                 // Check if line contains FOR token
                 IF FIND(IN1 := #lineBuffer.lines[#lineBuffer.pointers.retrievePointer].content, IN2 := #statKeyToken.tokenFor) <> 0 THEN
                   // Tokenize line where retrieve pointer is pointing at
                   #tempReturnVal := "LKinLang_TokenizeSlot"(lastIndexOfMerger := #statLastIndexOfMerger,
                                                             lineNumber := #lineBuffer.lines[#lineBuffer.pointers.retrievePointer].number,
                                                             line := #lineBuffer.lines[#lineBuffer.pointers.retrievePointer].content,
                                                             separators := #statSeparators,
                                                             mergers := #statMergers,
                                                             preprocessorConfig := #preProcessConfig,
                                                             tokenizedLine => #statTokenizedLine,
                                                             errorString := #statErrorString);

                   // Check if line has content
                   IF #statTokenizedLine.numberOfToken > 0 THEN
                     // Check if line starts with FOR token
                     IF #statTokenizedLine.lineToken[#statTokenizedLine.numberOfToken] = #statKeyToken.tokenFor THEN
                       // Increase array index
                       #statHierarchicLevel.numberOfLevels += 1;
                       // Check if index is ok
                       IF #statHierarchicLevel.numberOfLevels <= "LKINLANG_NUMBER_OF_HIERARCHICLEVEL" THEN
                         // Increase hierarchic level
                         #statHierarchicLevel.currentLevel += 1;
                         // Store entry
                         #statHierarchicLevel.levels[#statHierarchicLevel.numberOfLevels].level := #statHierarchicLevel.currentLevel;
                         #statHierarchicLevel.levels[#statHierarchicLevel.numberOfLevels].lineNumber := #statTokenizedLine.lineNo;
                         #statHierarchicLevel.levels[#statHierarchicLevel.numberOfLevels].type := "LKINLANG_ENTRY_TYPE_FOR"; // Type for FOR
                       ELSE
                         // Error hierarchic level array overflow
                         #statStatus := #ERR_HIERARCHIC_LEVEL_LIST;
                         #statStateIntern := #STATE_ERROR;
                         #statErrorString := CONCAT(IN1 := #statErrorString, IN2 := 'Error: Maximum array index of hierarchic level reached');
                         #statErrorString := CONCAT(IN1 := #statErrorString, IN2 := ' in line: ');
                         #statErrorString := CONCAT(IN1 := #statErrorString, IN2 := UDINT_TO_STRING(#statTokenizedLine.lineNo));
                       END_IF;
                     END_IF;
                   END_IF;
                 END_IF;

                 // Check if line contains ENDFOR token
                 IF FIND(IN1 := #lineBuffer.lines[#lineBuffer.pointers.retrievePointer].content, IN2 := #statKeyToken.tokenEndFor) <> 0 THEN
                   // Tokenize line where retrieve pointer is pointing at
                   #tempReturnVal := "LKinLang_TokenizeSlot"(lastIndexOfMerger := #statLastIndexOfMerger,
                                                             lineNumber := #lineBuffer.lines[#lineBuffer.pointers.retrievePointer].number,
                                                             line := #lineBuffer.lines[#lineBuffer.pointers.retrievePointer].content,
                                                             separators := #statSeparators,
                                                             mergers := #statMergers,
                                                             preprocessorConfig := #preProcessConfig,
                                                             tokenizedLine => #statTokenizedLine,
                                                             errorString := #statErrorString);

                   // Check if line has content
                   IF #statTokenizedLine.numberOfToken > 0 THEN
                     // Check if line starts with ENDFOR token
                     IF #statTokenizedLine.lineToken[#statTokenizedLine.numberOfToken] = #statKeyToken.tokenEndFor THEN
                       // Increase array index
                       #statHierarchicLevel.numberOfLevels += 1;
                       // Check if index is ok
                       IF #statHierarchicLevel.numberOfLevels <= "LKINLANG_NUMBER_OF_HIERARCHICLEVEL" THEN
                         // Store entry
                         #statHierarchicLevel.levels[#statHierarchicLevel.numberOfLevels].level := #statHierarchicLevel.currentLevel;
                         #statHierarchicLevel.levels[#statHierarchicLevel.numberOfLevels].lineNumber := #statTokenizedLine.lineNo;
                         #statHierarchicLevel.levels[#statHierarchicLevel.numberOfLevels].type := "LKINLANG_ENTRY_TYPE_ENDFOR"; // Type for ENDFOR

                         // Decrease hierarchic level
                         #statHierarchicLevel.currentLevel -= 1;
                       ELSE
                         // Error hierarchic level array overflow
                         #statStatus := #ERR_HIERARCHIC_LEVEL_LIST;
                         #statStateIntern := #STATE_ERROR;
                         #statErrorString := CONCAT(IN1 := #statErrorString, IN2 := 'Error: Maximum array index of hierarchic level reached');
                         #statErrorString := CONCAT(IN1 := #statErrorString, IN2 := ' in line: ');
                         #statErrorString := CONCAT(IN1 := #statErrorString, IN2 := UDINT_TO_STRING(#statTokenizedLine.lineNo));
                       END_IF;
                     END_IF;
                   END_IF;
                 END_IF;
               END_REGION GET_HIERARCHIC_LEVEL

               // Check if error occurred and exit reapeat
               IF #statStateIntern = #STATE_ERROR THEN
                 EXIT;
               END_IF;

               // ------------------------------------------------------------------------------------------
               // Search labels in program
               // ------------------------------------------------------------------------------------------
               // Check if LABEL key token is in line 
               // YES: Tokenize line
               // NO: next line
               REGION GENERATE_LABEL_LIST
                 // Check if line contains LABEL token
                 IF FIND(IN1 := #lineBuffer.lines[#lineBuffer.pointers.retrievePointer].content, IN2 := #statKeyToken.tokenJumpTarget) <> 0 THEN

                   // Tokenize line where retrieve pointer is pointing at
                   #tempReturnVal := "LKinLang_TokenizeSlot"(lastIndexOfMerger := #statLastIndexOfMerger,
                                                             lineNumber := #lineBuffer.lines[#lineBuffer.pointers.retrievePointer].number,
                                                             line := #lineBuffer.lines[#lineBuffer.pointers.retrievePointer].content,
                                                             separators := #statSeparators,
                                                             mergers := #statMergers,
                                                             preprocessorConfig := #preProcessConfig,
                                                             tokenizedLine => #statTokenizedLine,
                                                             errorString := #statErrorString);

                   // Check for error while tokenizing
                   IF #tempReturnVal <> 0 THEN
                     // Error while tokenizing
                     #statStatus := #ERR_TOKENIZING;
                     #statStateIntern := #STATE_ERROR;
                     EXIT;
                   END_IF;


                   // Check if line has content
                   IF #statTokenizedLine.numberOfToken > 0 THEN // Line has content --> Parse
                     // Go to ParseLine state if tokenizing was successful
                     // Check if line starts with 'LABEL'
                     IF #statTokenizedLine.lineToken[#statTokenizedLine.numberOfToken] = #statKeyToken.tokenJumpTarget THEN
                       // Check if line contains exactly 3 tokens
                       // Definition:
                       // [1] "myLabel"
                       // [2] " "
                       // [3] "LABEL"
                       IF #statTokenizedLine.numberOfToken = 3 THEN
                         IF #statTokenizedLine.lineToken[#statTokenizedLine.numberOfToken - 1] = ' ' // second token must be space
                           AND NOT "LKinLang_IsTokenNumberInclSign"(#statTokenizedLine.lineToken[#statTokenizedLine.numberOfToken - 2]) // first token must not be a number
                         THEN
                           // correct label definition 
                           // Check labelList if label already exists
                           FOR #tempCounter := 1 TO #statLabelList.numberOfLabels DO
                             IF #statLabelList.labels[#tempCounter].labelName = #statTokenizedLine.lineToken[#statTokenizedLine.numberOfToken - 2] THEN
                               // Label already exists in other line
                               // Throw error
                               #statStatus := #ERR_LABEL_LIST;
                               #statStateIntern := #STATE_ERROR;
                               #statErrorString := CONCAT(IN1 := #statErrorString, IN2 := ';Error: Label is not unique');
                               #statErrorString := CONCAT(IN1 := #statErrorString, IN2 := ' in line: ');
                               #statErrorString := CONCAT(IN1 := #statErrorString, IN2 := UDINT_TO_STRING(#statTokenizedLine.lineNo));
                               EXIT;
                             END_IF;
                           END_FOR;

                           // Check if error was set in for loop
                           // --> Abort repeat loop 
                           IF #statStateIntern = #STATE_ERROR THEN
                             EXIT;
                           END_IF;

                           // Check if name is a keyword
                           IF "LKinLang_IsTokenKeyWord"(token := #statTokenizedLine.lineToken[#statTokenizedLine.numberOfToken - 2], keyToken := #statKeyToken) THEN
                             // Error: Label name can not be a keyword
                             #statStatus := #ERR_LABEL_LIST;
                             #statStateIntern := #STATE_ERROR;
                             #statErrorString := CONCAT(IN1 := #statErrorString, IN2 := 'Error: Label name must not be a keyword');
                             #statErrorString := CONCAT(IN1 := #statErrorString, IN2 := '; Line: ');
                             #statErrorString := CONCAT(IN1 := #statErrorString, IN2 := UDINT_TO_STRING(#statTokenizedLine.lineNo));
                             EXIT;
                           END_IF;

                           // Check if name is a parameter 
                           FOR #tempVarIndex := 1 TO "LKINLANG_MAX_NUMBER_OF_PARAMETERS" DO
                             IF #statParameterLookUpTable[#tempVarIndex].parameterNameString = #statTokenizedLine.lineToken[#statTokenizedLine.numberOfToken - 2] THEN
                               // Error: Label name can not be a parameter
                               #statStatus := #ERR_LABEL_LIST;
                               #statStateIntern := #STATE_ERROR;
                               #statErrorString := CONCAT(IN1 := #statErrorString, IN2 := 'Error: Label name must not be a keyword');
                               #statErrorString := CONCAT(IN1 := #statErrorString, IN2 := '; Line: ');
                               #statErrorString := CONCAT(IN1 := #statErrorString, IN2 := UDINT_TO_STRING(#statTokenizedLine.lineNo));
                               EXIT;
                             END_IF;
                           END_FOR;

                           // Check if error was set in for loop
                           // --> Abort repeat loop 
                           IF #statStateIntern = #STATE_ERROR THEN
                             EXIT;
                           END_IF;

                           // Check if the number of labels is ok 
                           IF #statLabelList.numberOfLabels >= "LKINLANG_NUMBER_OF_LABELS" THEN
                             // No more space in labelList
                             // Throw error 
                             #statStatus := #ERR_LABEL_LIST;
                             #statStateIntern := #STATE_ERROR;
                             #statErrorString := CONCAT(IN1 := #statErrorString, IN2 := ';Error: Maximum number of labels reached');
                             #statErrorString := CONCAT(IN1 := #statErrorString, IN2 := ' in line: ');
                             #statErrorString := CONCAT(IN1 := #statErrorString, IN2 := UDINT_TO_STRING(#statTokenizedLine.lineNo));
                             EXIT;
                           END_IF;

                           IF #statStateIntern <> #STATE_ERROR THEN
                             // Increment number of labels
                             #statLabelList.numberOfLabels += 1;
                             // Set the label info
                             #statLabelList.labels[#statLabelList.numberOfLabels].labelName := #statTokenizedLine.lineToken[#statTokenizedLine.numberOfToken - 2];
                             #statLabelList.labels[#statLabelList.numberOfLabels].lineNumber := #statTokenizedLine.lineNo;
                             IF #statHierarchicLevel.numberOfLevels > 0 THEN
                               #statLabelList.labels[#statLabelList.numberOfLabels].hierarchicLevel := #statHierarchicLevel.levels[#statHierarchicLevel.numberOfLevels].level;
                             ELSE
                               #statLabelList.labels[#statLabelList.numberOfLabels].hierarchicLevel := 0;
                             END_IF;
                           ELSE
                             // Error was set already set
                             // Do nothing
                             ;
                           END_IF;

                         ELSE
                           // Wrong label definition --> No space or correct name
                           // Throw error
                           #statStatus := #ERR_LABEL_LIST;
                           #statStateIntern := #STATE_ERROR;
                           #statErrorString := CONCAT(IN1 := #statErrorString, IN2 := ';Error: Invalid label definition');
                           #statErrorString := CONCAT(IN1 := #statErrorString, IN2 := ' in line: ');
                           #statErrorString := CONCAT(IN1 := #statErrorString, IN2 := UDINT_TO_STRING(#statTokenizedLine.lineNo));
                           EXIT;
                         END_IF;
                       ELSE
                         // Wrong label definition --> Not 3 token
                         // Throw error
                         #statStatus := #ERR_LABEL_LIST;
                         #statStateIntern := #STATE_ERROR;
                         #statErrorString := CONCAT(IN1 := #statErrorString, IN2 := ';Error: Invalid label definition');
                         #statErrorString := CONCAT(IN1 := #statErrorString, IN2 := ' in line: ');
                         #statErrorString := CONCAT(IN1 := #statErrorString, IN2 := UDINT_TO_STRING(#statTokenizedLine.lineNo));
                         EXIT;
                       END_IF;

                     ELSE
                       ;// Not a label definition
                     END_IF;
                   ELSE
                     ; // Line is empty --> Tokenize next Line
                   END_IF;
                 END_IF;
               END_REGION GENERATE_LABEL_LIST

               // ------------------------------------------------------------------------------------------
               // Search sub programs
               // ------------------------------------------------------------------------------------------
               // Check if SUB key token is in line 
               REGION SUB_PROGRAM
                 // Check if line contains SUB token
                 IF FIND(IN1 := #lineBuffer.lines[#lineBuffer.pointers.retrievePointer].content, IN2 := #statKeyToken.tokenStartSub) <> 0 THEN

                   // Tokenize line where retrieve pointer is pointing at
                   #tempReturnVal := "LKinLang_TokenizeSlot"(lastIndexOfMerger := #statLastIndexOfMerger,
                                                             lineNumber := #lineBuffer.lines[#lineBuffer.pointers.retrievePointer].number,
                                                             line := #lineBuffer.lines[#lineBuffer.pointers.retrievePointer].content,
                                                             separators := #statSeparators,
                                                             mergers := #statMergers,
                                                             preprocessorConfig := #preProcessConfig,
                                                             tokenizedLine => #statTokenizedLine,
                                                             errorString := #statErrorString);

                   // Check for error while tokenizing
                   IF #tempReturnVal <> 0 THEN
                     // Error while tokenizing
                     #statStatus := #ERR_TOKENIZING;
                     #statStateIntern := #STATE_ERROR;
                     EXIT;
                   END_IF;

                   // Check if line has content
                   IF #statTokenizedLine.numberOfToken > 0 THEN // Line has content --> Parse
                     // Check if line starts with 'SUB'
                     IF #statTokenizedLine.lineToken[#statTokenizedLine.numberOfToken] = #statKeyToken.tokenStartSub THEN
                       // Check if line contains exactly 3 tokens
                       // Definition:
                       // [1] "mySubPrg_1"
                       // [2] " "
                       // [3] "SUB"
                       IF #statTokenizedLine.numberOfToken = 3 THEN
                         IF #statTokenizedLine.lineToken[#statTokenizedLine.numberOfToken - 1] = ' ' // second token must be space
                           AND NOT "LKinLang_IsTokenNumberInclSign"(#statTokenizedLine.lineToken[#statTokenizedLine.numberOfToken - 2]) // first token must not be a number
                         THEN
                           // correct sub definition 
                           // Check subPrgList if sub already exists
                           FOR #tempCounter := 1 TO #statSubPrgList.numberOfSubPrgs DO
                             IF #statSubPrgList.subPrgs[#tempCounter].prgName = #statTokenizedLine.lineToken[#statTokenizedLine.numberOfToken - 2] THEN
                               // Sub already exists in other line
                               // Throw error
                               #statStatus := #ERR_SUB_PROGRAM_LIST;
                               #statStateIntern := #STATE_ERROR;
                               #statErrorString := CONCAT(IN1 := #statErrorString, IN2 := ';Error: Subprogram is not unique');
                               #statErrorString := CONCAT(IN1 := #statErrorString, IN2 := ' in line: ');
                               #statErrorString := CONCAT(IN1 := #statErrorString, IN2 := UDINT_TO_STRING(#statTokenizedLine.lineNo));
                               EXIT;
                             END_IF;
                           END_FOR;

                           // Check if error was set in for loop
                           // --> Abort repeat loop 
                           IF #statStateIntern = #STATE_ERROR THEN
                             EXIT;
                           END_IF;

                           // Check if name is a keyword
                           IF "LKinLang_IsTokenKeyWord"(token := #statTokenizedLine.lineToken[#statTokenizedLine.numberOfToken - 2], keyToken := #statKeyToken) THEN
                             // Error: Variable name can not be a keyword
                             #statStatus := #ERR_SUB_PROGRAM_LIST;
                             #statStateIntern := #STATE_ERROR;
                             #statErrorString := CONCAT(IN1 := #statErrorString, IN2 := 'Error: Subprogram name must not be a keyword');
                             #statErrorString := CONCAT(IN1 := #statErrorString, IN2 := '; Line: ');
                             #statErrorString := CONCAT(IN1 := #statErrorString, IN2 := UDINT_TO_STRING(#statTokenizedLine.lineNo));
                             EXIT;
                           END_IF;

                           // Check if name is a parameter 
                           FOR #tempVarIndex := 1 TO "LKINLANG_MAX_NUMBER_OF_PARAMETERS" DO
                             IF #statParameterLookUpTable[#tempVarIndex].parameterNameString = #statTokenizedLine.lineToken[#statTokenizedLine.numberOfToken - 2] THEN
                               // Error: Variable name can not be a keyword
                               #statStatus := #ERR_SUB_PROGRAM_LIST;
                               #statStateIntern := #STATE_ERROR;
                               #statErrorString := CONCAT(IN1 := #statErrorString, IN2 := 'Error: Subprogram name must not be a keyword');
                               #statErrorString := CONCAT(IN1 := #statErrorString, IN2 := '; Line: ');
                               #statErrorString := CONCAT(IN1 := #statErrorString, IN2 := UDINT_TO_STRING(#statTokenizedLine.lineNo));
                               EXIT;
                             END_IF;
                           END_FOR;

                           // Check if error was set in for loop
                           // --> Abort repeat loop 
                           IF #statStateIntern = #STATE_ERROR THEN
                             EXIT;
                           END_IF;

                           // Check if the number of labels is ok 
                           IF #statSubPrgList.numberOfSubPrgs >= "LKINLANG_NUMBER_OF_SUBPROGRAMS" THEN
                             // No more space in subPrgList
                             // Throw error 
                             #statStatus := #ERR_SUB_PROGRAM_LIST;
                             #statStateIntern := #STATE_ERROR;
                             #statErrorString := CONCAT(IN1 := #statErrorString, IN2 := ';Error: Maximum number of subprograms reached');
                             #statErrorString := CONCAT(IN1 := #statErrorString, IN2 := ' in line: ');
                             #statErrorString := CONCAT(IN1 := #statErrorString, IN2 := UDINT_TO_STRING(#statTokenizedLine.lineNo));
                             EXIT;
                           END_IF;

                           IF #statStateIntern <> #STATE_ERROR THEN
                             // Increment number of labels
                             #statSubPrgList.numberOfSubPrgs += 1;
                             // Set the label info
                             #statSubPrgList.subPrgs[#statSubPrgList.numberOfSubPrgs].prgName := #statTokenizedLine.lineToken[#statTokenizedLine.numberOfToken - 2];
                             #statSubPrgList.subPrgs[#statSubPrgList.numberOfSubPrgs].lineNumberStart := #statTokenizedLine.lineNo;
                           ELSE
                             // Error was set already set
                             // Do nothing
                             ;
                           END_IF;

                         ELSE
                           // Wrong label definition --> No space or correct name
                           // Throw error
                           #statStatus := #ERR_SUB_PROGRAM_LIST;
                           #statStateIntern := #STATE_ERROR;
                           #statErrorString := CONCAT(IN1 := #statErrorString, IN2 := ';Error: Invalid subprogram definition');
                           #statErrorString := CONCAT(IN1 := #statErrorString, IN2 := ' in line: ');
                           #statErrorString := CONCAT(IN1 := #statErrorString, IN2 := UDINT_TO_STRING(#statTokenizedLine.lineNo));
                           EXIT;
                         END_IF;
                       ELSE
                         // Wrong label definition --> Not 3 token
                         // Throw error
                         #statStatus := #ERR_SUB_PROGRAM_LIST;
                         #statStateIntern := #STATE_ERROR;
                         #statErrorString := CONCAT(IN1 := #statErrorString, IN2 := ';Error: Invalid subprogram definition');
                         #statErrorString := CONCAT(IN1 := #statErrorString, IN2 := ' in line: ');
                         #statErrorString := CONCAT(IN1 := #statErrorString, IN2 := UDINT_TO_STRING(#statTokenizedLine.lineNo));
                         EXIT;
                       END_IF;
                     ELSE
                       ; // Does not start with key token
                     END_IF;
                   ELSE
                     ; // Empty line
                   END_IF;
                 END_IF;

                 // Check if line contains END SUB token
                 IF FIND(IN1 := #lineBuffer.lines[#lineBuffer.pointers.retrievePointer].content, IN2 := #statKeyToken.tokenEndSub) <> 0 THEN
                   // Tokenize line where retrieve pointer is pointing at
                   #tempReturnVal := "LKinLang_TokenizeSlot"(lastIndexOfMerger := #statLastIndexOfMerger,
                                                             lineNumber := #lineBuffer.lines[#lineBuffer.pointers.retrievePointer].number,
                                                             line := #lineBuffer.lines[#lineBuffer.pointers.retrievePointer].content,
                                                             separators := #statSeparators,
                                                             mergers := #statMergers,
                                                             preprocessorConfig := #preProcessConfig,
                                                             tokenizedLine => #statTokenizedLine,
                                                             errorString := #statErrorString);

                   // Check for error while tokenizing
                   IF #tempReturnVal <> 0 THEN
                     // Error while tokenizing
                     #statStatus := #ERR_TOKENIZING;
                     #statStateIntern := #STATE_ERROR;
                     EXIT;
                   END_IF;

                   // Check if line has content
                   IF #statTokenizedLine.numberOfToken > 0 THEN
                     IF #statTokenizedLine.numberOfToken = 2 THEN
                       IF CONCAT(IN1 := #statTokenizedLine.lineToken[#statTokenizedLine.numberOfToken], IN2 := #statTokenizedLine.lineToken[#statTokenizedLine.numberOfToken - 1]) <> #statKeyToken.tokenEndSub THEN
                         // Throw error
                         #statStatus := #ERR_SUB_PROGRAM_LIST;
                         #statStateIntern := #STATE_ERROR;
                         #statErrorString := CONCAT(IN1 := #statErrorString, IN2 := ';Error: Invalid end of subprogram definition');
                         #statErrorString := CONCAT(IN1 := #statErrorString, IN2 := ' in line: ');
                         #statErrorString := CONCAT(IN1 := #statErrorString, IN2 := UDINT_TO_STRING(#statTokenizedLine.lineNo));
                         EXIT;
                       END_IF;
                     ELSIF #statTokenizedLine.numberOfToken = 1 THEN
                       IF #statTokenizedLine.lineToken[#statTokenizedLine.numberOfToken] <> #statKeyToken.tokenEndSub THEN
                         // Throw error
                         #statStatus := #ERR_SUB_PROGRAM_LIST;
                         #statStateIntern := #STATE_ERROR;
                         #statErrorString := CONCAT(IN1 := #statErrorString, IN2 := ';Error: Invalid end of subprogram definition');
                         #statErrorString := CONCAT(IN1 := #statErrorString, IN2 := ' in line: ');
                         #statErrorString := CONCAT(IN1 := #statErrorString, IN2 := UDINT_TO_STRING(#statTokenizedLine.lineNo));
                         EXIT;
                       END_IF;
                     ELSE
                       // Throw error
                       #statStatus := #ERR_SUB_PROGRAM_LIST;
                       #statStateIntern := #STATE_ERROR;
                       #statErrorString := CONCAT(IN1 := #statErrorString, IN2 := ';Error: Invalid end of subprogram definition');
                       #statErrorString := CONCAT(IN1 := #statErrorString, IN2 := ' in line: ');
                       #statErrorString := CONCAT(IN1 := #statErrorString, IN2 := UDINT_TO_STRING(#statTokenizedLine.lineNo));
                       EXIT;
                     END_IF;

                     // Check if definition was ok
                     IF #statStateIntern <> #STATE_ERROR THEN
                       // Check if end of sub program is allowed 
                       IF #statSubPrgList.subPrgs[#statSubPrgList.numberOfSubPrgs].lineNumberEnd = 0 THEN
                         ; // OK store linenumber
                         #statSubPrgList.subPrgs[#statSubPrgList.numberOfSubPrgs].lineNumberEnd := #statTokenizedLine.lineNo;
                       ELSE
                         ; // end was already set --> error?
                         // Throw error
                         #statStatus := #ERR_SUB_PROGRAM_LIST;
                         #statStateIntern := #STATE_ERROR;
                         #statErrorString := CONCAT(IN1 := #statErrorString, IN2 := ';Error: Invalid end of subprogram');
                         #statErrorString := CONCAT(IN1 := #statErrorString, IN2 := ' in line: ');
                         #statErrorString := CONCAT(IN1 := #statErrorString, IN2 := UDINT_TO_STRING(#statTokenizedLine.lineNo));
                         EXIT;
                       END_IF;
                     END_IF;

                   ELSE
                     ; // Empty line
                   END_IF;
                 END_IF;

               END_REGION SUB_PROGRAM

               // Check if error occurred and exit reapeat
               IF #statStateIntern = #STATE_ERROR THEN
                 EXIT;
               END_IF;

               // Increase line counter --> Count every line; not just empty ones
               #tempEmptyLineCounter += 1;

               // Check empty line counter to abort repeat
               IF #tempEmptyLineCounter >= #MAX_LINES_LABEL_LIST THEN
                 #tempAbortRepeat := TRUE;
               END_IF;

             ELSE
               // Waiting for line buffer --> do nothing
               // Abort repeat
               #tempAbortRepeat := TRUE;
             END_IF;

             // Check if end of file was reached --> Set by FileHandler
             // YES: Abort this repeat and restart fileHandler to read lines from start again
             // NO: Continue with label list
             IF #lineBuffer.pointers.endOfFile
               AND #lineBuffer.pointers.addPointer = #lineBuffer.pointers.retrievePointer
             THEN
               // Check if the line number is greater the retireve Pointer --> If yes then a buffer overflow occured and restart is neccessary
               IF #lineBuffer.lines[#lineBuffer.pointers.retrievePointer].number > #lineBuffer.pointers.retrievePointer THEN
                 #lineBuffer.pointers.restart := TRUE;
               END_IF;
               #lineBuffer.pointers.retrievePointer := 0;
               #statFBState := #FB_STATE_PARSING;
               #tempAbortRepeat := TRUE;

             ELSIF #lineBuffer.pointers.ignoreAddPointer AND #lineBuffer.pointers.retrievePointer > 0 THEN
               IF #lineBuffer.lines[#lineBuffer.pointers.retrievePointer].number = 0 THEN
                 #lineBuffer.pointers.retrievePointer := 0;
                 #statFBState := #FB_STATE_PARSING;
                 #tempAbortRepeat := TRUE;
               END_IF;
             END_IF;

           UNTIL #tempAbortRepeat END_REPEAT;

           // Check if found subprgs are ok 
           IF #statFBState = #FB_STATE_PARSING THEN // Signalizes that precheck is done
             FOR #tempCounter := 1 TO #statSubPrgList.numberOfSubPrgs DO
               IF #statSubPrgList.subPrgs[#tempCounter].lineNumberStart = 0 THEN
                 // Throw error
                 #statStatus := #ERR_SUB_PROGRAM_LIST;
                 #statStateIntern := #STATE_ERROR;
                 #statErrorString := CONCAT(IN1 := #statErrorString, IN2 := 'Error: Missing start of subprogram');
                 EXIT;
               END_IF;
               IF #statSubPrgList.subPrgs[#tempCounter].lineNumberEnd = 0 THEN
                 // Throw error
                 #statStatus := #ERR_SUB_PROGRAM_LIST;
                 #statStateIntern := #STATE_ERROR;
                 #statErrorString := CONCAT(IN1 := #statErrorString, IN2 := 'Error: Missing end of subprogram started in line: ');
                 #statErrorString := CONCAT(IN1 := #statErrorString, IN2 := UDINT_TO_STRING(#statSubPrgList.subPrgs[#tempCounter].lineNumberStart));
                 EXIT;
               END_IF;
             END_FOR;
           END_IF;

           // ------------------------------------------------------------------------------------------
           // Error state for internal case
           // Switch to in case of error and do not execute other states
           // ------------------------------------------------------------------------------------------ 
           REGION ERROR_STATE
             // Error State 
             IF #statStateIntern = #STATE_ERROR THEN
               // Reset lineBuffer pointer
               #lineBuffer.pointers.retrievePointer := 0;
               #lineBuffer.pointers.addPointerRestarted := FALSE;
               // Reset file state
               IF #lineBuffer.info.fileState = "LKINLANG_FILE_STATE_RUNNING" THEN
                 #lineBuffer.info.fileState := "LKINLANG_FILE_STATE_IDLE";
               END_IF;
             END_IF;
           END_REGION ERROR_STATE
         END_REGION FB_STATE_PRECHECK_PRG

         // ------------------------------------------------------------------------------------------
         // Main routine of FB
         // Activated after init steps are done 
         // Works with internal states (IF cases) to parse and write one line/cmd per cycle
         // ------------------------------------------------------------------------------------------ 
       #FB_STATE_PARSING: // Parsing active
         REGION FB_STATE_PARSING
           // For loop to process more lines in one OB cycle
           FOR #tempCycleCounter := 1 TO #MAX_LINES_PER_CYCLE DO

             // ------------------------------------------------------------------------------------------
             // Search line
             // Check if searched line is already in lineBuffer
             // YES: Go to STATE_TOKENIZING
             // NO: Go to STATE_FILEHANDLER_REQUEST
             // ------------------------------------------------------------------------------------------ 
             REGION SEARCH_LINE
               IF #statStateIntern = #STATE_SEARCH_LINE THEN
                 // ----------------------------
                 // Search if line is in lineBuffer already
                 // ----------------------------
                 #tempConditionResult := FALSE;
                 FOR #tempCounter := "LKINLANG_FIRST_INDEX_LINE_BUFFER" TO "LKINLANG_LAST_INDEX_LINE_BUFFER" DO
                   IF #lineBuffer.lines[#tempCounter].number = #statSearchedLine THEN
                     #tempConditionResult := TRUE;// Line was found
                     EXIT;
                   ELSE
                     CONTINUE;
                   END_IF;
                 END_FOR;

                 IF #tempConditionResult = FALSE THEN
                   // ----------------------------
                   // Line is not in lineBuffer
                   // --> Request from fileHandler
                   // ----------------------------
                   #lineBuffer.pointers.requestedLine := #statSearchedLine;
                   // Restart FileHandler if necessary
                   IF #lineBuffer.pointers.endOfFile THEN
                     #lineBuffer.pointers.restart := TRUE;
                   END_IF;

                   // Go to next state
                   #statStateIntern := #STATE_FILEHANDLER_REQUEST;

                 ELSE
                   // ----------------------------
                   // Line is in lineBuffer
                   // ----------------------------
                   #lineBuffer.pointers.retrievePointer := #tempCounter; // Set retrievePointer to line in lineBuffer

                   // Set / Reset "addPointerRestarted"
                   IF #lineBuffer.pointers.addPointerRestarted = TRUE
                     AND #tempCounter <= #lineBuffer.pointers.addPointer
                   THEN
                     #lineBuffer.pointers.addPointerRestarted := FALSE;

                   ELSIF #lineBuffer.pointers.addPointerRestarted = FALSE
                     AND #tempCounter > #lineBuffer.pointers.addPointer
                   THEN
                     #lineBuffer.pointers.addPointerRestarted := TRUE;
                   END_IF;

                   // Go to next state
                   #statStateIntern := #STATE_TOKENIZING;
                 END_IF;
               END_IF;
             END_REGION SEARCH_LINE

             // ------------------------------------------------------------------------------------------
             // FILEHANDLER_REQUEST
             // Searched line was requested from fileHandler, check if available
             // YES: Go to STATE_TOKENIZING
             // NO: Wait here
             // ------------------------------------------------------------------------------------------ 
             REGION FILEHANDLER_REQUEST
               IF #statStateIntern = #STATE_FILEHANDLER_REQUEST THEN
                 // Check if fileHandler has found the line
                 IF #lineBuffer.pointers.addPointer <> 0
                   AND #lineBuffer.pointers.retrievePointer = 0
                   AND #lineBuffer.pointers.addPointerRestarted = FALSE
                 THEN
                   // Line found --> Set retrieve pointer to written index
                   #lineBuffer.pointers.retrievePointer := #lineBuffer.pointers.addPointer;
                   #statStateIntern := #STATE_TOKENIZING;
                 ELSE
                   ; // Wait in this state
                 END_IF;
               END_IF;
             END_REGION FILEHANDLER_REQUEST

             // ------------------------------------------------------------------------------------------
             // Tokenize line
             // Check pointers and increase retrieve pointer
             // Get line from buffer and tokenize it
             // Go to Parse_Line state
             // ------------------------------------------------------------------------------------------ 
             REGION TOKENIZE_LINE
               // Tokenize line
               IF #statStateIntern = #STATE_TOKENIZING
               THEN

                 // Reset empty line counter
                 #tempEmptyLineCounter := 0;

                 // Repeat tokenizing until aborted
                 // Aborted by:
                 // - Line with content
                 // - Empty line counter higher as MAX_EMPTY_LINES_PER_CYCLE
                 // - No more lines in line buffer
                 REPEAT

                   #tempPointerOk := FALSE; // Init temp

                   IF #lineBuffer.pointers.ignoreAddPointer THEN
                     #tempPointerOk := TRUE;
                   ELSIF #lineBuffer.pointers.bufferLocked THEN
                     #tempPointerOk := FALSE;
                   ELSIF #statSearchedLine <> 0 THEN
                     #tempPointerOk := TRUE;
                   ELSIF #lineBuffer.pointers.addPointerRestarted = FALSE THEN
                     #tempPointerOk := #lineBuffer.pointers.addPointer > #lineBuffer.pointers.retrievePointer;
                   ELSIF #lineBuffer.pointers.addPointerRestarted = TRUE THEN
                     #tempPointerOk := #lineBuffer.pointers.addPointer < #lineBuffer.pointers.retrievePointer;
                   END_IF;

                   // Check lineBuffer pointer if next line can be retrieved
                   // IF ((#lineBuffer.pointers.addPointer > #lineBuffer.pointers.retrievePointer
                   //   AND NOT #lineBuffer.pointers.bufferLocked // Buffer is not locked by fileHandler
                   //   AND NOT #lineBuffer.pointers.addPointerRestarted) // Overflow of ring buffer
                   //   OR
                   //   (#lineBuffer.pointers.addPointer < #lineBuffer.pointers.retrievePointer
                   //   AND #lineBuffer.pointers.addPointerRestarted
                   //   AND NOT #lineBuffer.pointers.bufferLocked))
                   //   OR #lineBuffer.pointers.ignoreAddPointer // FR 25.11.2019
                   // THEN
                   IF #tempPointerOk THEN
                     IF #statSearchedLine <= 0 THEN
                       // Increment retrieve pointer
                       IF #lineBuffer.pointers.retrievePointer < "LKINLANG_LAST_INDEX_LINE_BUFFER" THEN
                         #lineBuffer.pointers.retrievePointer += 1;

                         // Reset retrieve pointer to 1 and reset overflow variable
                       ELSIF #lineBuffer.pointers.retrievePointer >= "LKINLANG_LAST_INDEX_LINE_BUFFER" THEN
                         #lineBuffer.pointers.retrievePointer := 1;
                         #lineBuffer.pointers.addPointerRestarted := FALSE;
                       END_IF;
                     ELSE
                       // Line was searched
                       // -> Reset static
                       // -> Do not change pointer as they were already set before
                       #statSearchedLine := 0;
                     END_IF;

                     // Tokenize line where retrieve pointer is pointing at
                     #tempReturnVal := "LKinLang_TokenizeSlot"(lastIndexOfMerger := #statLastIndexOfMerger,
                                                               lineNumber := #lineBuffer.lines[#lineBuffer.pointers.retrievePointer].number,
                                                               line := #lineBuffer.lines[#lineBuffer.pointers.retrievePointer].content,
                                                               separators := #statSeparators,
                                                               mergers := #statMergers,
                                                               preprocessorConfig := #preProcessConfig,
                                                               tokenizedLine => #statTokenizedLine,
                                                               errorString := #statErrorString);

                     // Check for error while tokenizing
                     IF #tempReturnVal <> 0 THEN
                       // Error while tokenizing
                       #statStatus := #ERR_TOKENIZING;
                       #statStateIntern := #STATE_ERROR;
                       EXIT;
                     END_IF;

                     // Check if line has content
                     IF #statTokenizedLine.numberOfToken > 0 THEN // Line has content --> Parse
                       // Go to ParseLine state if tokenizing was successful
                       #statStateIntern := #STATE_INIT_PARSE_LINE;

                       // Abort repeat
                       #tempAbortRepeat := TRUE;
                     ELSE
                       // Line is empty --> Tokenize next Line
                       #tempEmptyLineCounter += 1;

                       IF #lineBuffer.pointers.ignoreAddPointer
                         AND #lineBuffer.pointers.retrievePointer = "LKINLANG_LAST_INDEX_LINE_BUFFER" THEN
                         // Error no more lines but haven't found endOfPrg (M30) yet
                         // Throw error
                         #statStatus := #ERR_PARSING;
                         #statStateIntern := #STATE_ERROR;
                         #statErrorString := CONCAT(IN1 := #statErrorString, IN2 := 'Error: Missing end of program(M30) or subprogram(ENDSUB) in line ');
                         #statErrorString := CONCAT(IN1 := #statErrorString, IN2 := UDINT_TO_STRING(#statTokenizedLine.lineNo));
                         EXIT;
                       END_IF;

                     END_IF;

                     IF #tempEmptyLineCounter >= #MAX_EMPTY_LINES_PER_CYCLE THEN
                       #tempAbortRepeat := TRUE;
                     END_IF;

                   ELSE
                     // Waiting for line buffer --> do nothing
                     // Abort repeat
                     #tempAbortRepeat := TRUE;

                     IF #lineBuffer.pointers.endOfFile
                       AND #lineBuffer.pointers.addPointer = #lineBuffer.pointers.retrievePointer
                     THEN
                       // Error no more lines but haven't found endOfPrg (M30) yet
                       // Throw error
                       #statStatus := #ERR_PARSING;
                       #statStateIntern := #STATE_ERROR;
                       #statErrorString := CONCAT(IN1 := #statErrorString, IN2 := 'Error: Missing end of program(M30) or subprogram(ENDSUB) in line ');
                       #statErrorString := CONCAT(IN1 := #statErrorString, IN2 := UDINT_TO_STRING(#statTokenizedLine.lineNo));
                       EXIT;
                     END_IF;
                   END_IF;

                 UNTIL #tempAbortRepeat END_REPEAT;

               END_IF;
             END_REGION TOKENIZE_LINE

             // ------------------------------------------------------------------------------------------
             // Init parse line
             // Initialize parsing of line
             // Go to IS_LINE_VARIABLE_DEFINITION state
             // ------------------------------------------------------------------------------------------ 
             REGION INIT_PARSE_LINE
               // Initialize varaibles for parsing one line
               IF #statStateIntern = #STATE_INIT_PARSE_LINE
               THEN
                 // Init token counter
                 #tempTokenCounter := 1;

                 // Init condition counter
                 #tempConditionCounter := 1;

                 #statRightSideOfEquation := TRUE;
                 #statStringExpression := '';

                 // Init element in line counter
                 #statElementCounterInLine := #statElementCounterEmpty;

                 // Init parameter counter in line
                 FOR #tempCounter := 1 TO "LKINLANG_NUMBER_OF_CONDITIONS" DO
                   #statSetParametersInLine[#tempCounter] := #statConditionEmpty;
                 END_FOR;

                 // Initialize actual command
                 #statActualCommand := #statPathDataElementEmpty;

                 // Reset parameter valid bits --> They are set to TRUE when the coordinate was parsed
                 FOR #tempCounter := 1 TO "LKINCTRL_NO_OF_VALID_BITS" DO
                   #statActualCommand.pathDataElement.parameterValid[#tempCounter] := FALSE;
                 END_FOR;

                 // testing FR 2019.03.12
                 // Reset condition for check in line
                 FOR #tempCounter := 1 TO "LKINLANG_NUMBER_OF_CONDITIONS" DO
                   IF #statConditionsToCheck[#tempCounter].Mode = "LKINLANG_CONDITION_IN_LINE" THEN
                     #statConditionsToCheck[#tempCounter] := #statConditionEmpty;
                   END_IF;
                 END_FOR;

                 // Next step 
                 #statStateIntern := #STATE_IS_LINE_VAR_DEF;
               END_IF;
             END_REGION INIT_PARSE_LINE


             // ------------------------------------------------------------------------------------------
             // Is line variable definition
             // Check if the line contains a variable definition like "DEF DINT myVar_1"
             // YES: Go to STATE_LINE_IS_VAR_DEF
             // NO: Go to IS_LINE_LABEL 
             // ------------------------------------------------------------------------------------------ 
             REGION IS_LINE_VARIABLE_DEFINITION
               IF #statStateIntern = #STATE_IS_LINE_VAR_DEF
               THEN
                 // Check if line contains variable definition 
                 // YES: Create variable
                 // NO: Continue with normal check